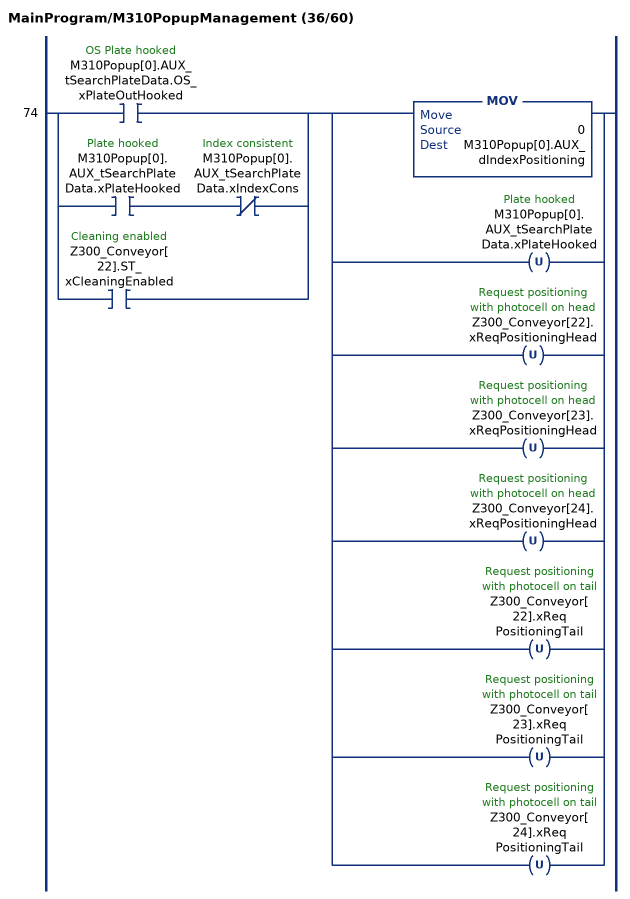
   74: [XIC(M310Popup[0].AUX_tSearchPlateData.OS_xPlateOutHooked) ,XIC(M310Popup[0].AUX_tSearchPlateData.xPlateHooked) XIO(M310Popup[0].AUX_tSearchPlateData.xIndexCons) ,XIC(Z300_Conveyor[22].ST_xCleaningEnabled) ][MOV(0,M310Popup[0].AUX_dIndexPositioning) ,OTU(M310Popup[0].AUX_tSearchPlateData.xPlateHooked) ,OTU(Z300_Conveyor[22].xReqPositioningHead) ,OTU(Z300_Conveyor[23].xReqPositioningHead) ,OTU(Z300_Conveyor[24].xReqPositioningHead) ,OTU(Z300_Conveyor[22].xReqPositioningTail) ,OTU(Z300_Conveyor[23].xReqPositioningTail) ,OTU(Z300_Conveyor[24].xReqPositioningTail) ];
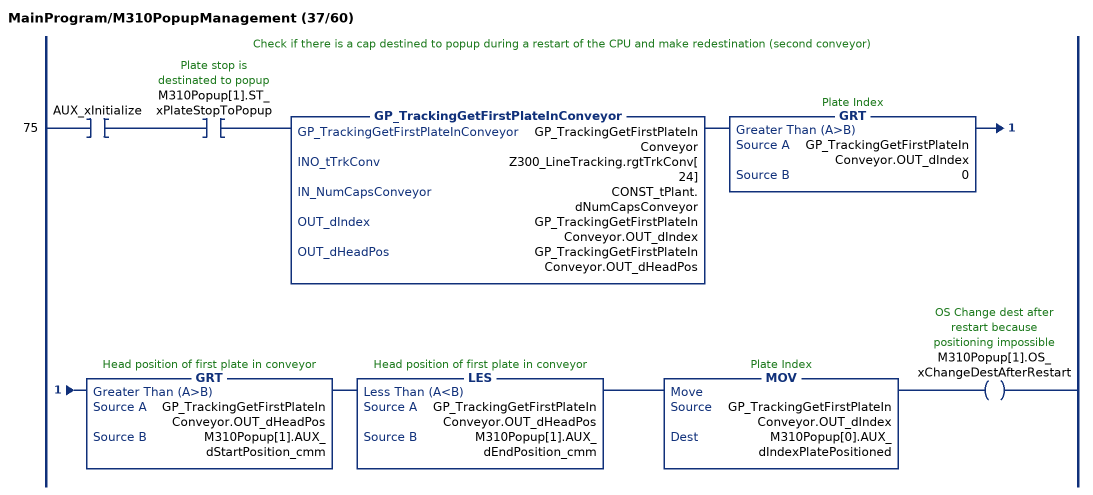
   // Check if there is a cap destined to popup during a restart of the CPU and make redestination (second conveyor)
   75: XIC(AUX_xInitialize)XIC(M310Popup[1].ST_xPlateStopToPopup)GP_TrackingGetFirstPlateInConveyor(GP_TrackingGetFirstPlateInConveyor,Z300_LineTracking.rgtTrkConv[24],CONST_tPlant.dNumCapsConveyor,GP_TrackingGetFirstPlateInConveyor.OUT_dIndex,GP_TrackingGetFirstPlateInConveyor.OUT_dHeadPos)GRT(GP_TrackingGetFirstPlateInConveyor.OUT_dIndex,0)GRT(GP_TrackingGetFirstPlateInConveyor.OUT_dHeadPos,M310Popup[1].AUX_dStartPosition_cmm)LES(GP_TrackingGetFirstPlateInConveyor.OUT_dHeadPos,M310Popup[1].AUX_dEndPosition_cmm)MOV(GP_TrackingGetFirstPlateInConveyor.OUT_dIndex,M310Popup[0].AUX_dIndexPlatePositioned)OTE(M310Popup[1].OS_xChangeDestAfterRestart);
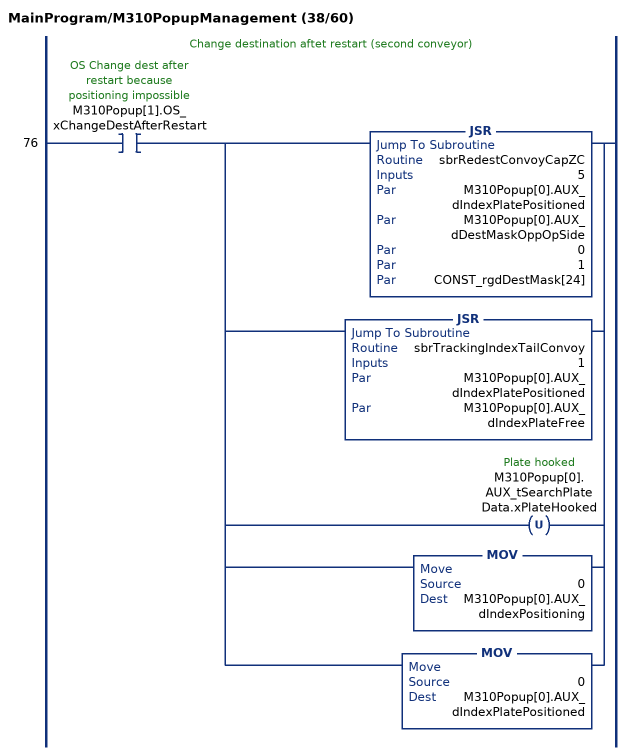
   // Change destination aftet restart (second conveyor)
   76: XIC(M310Popup[1].OS_xChangeDestAfterRestart)[JSR(sbrRedestConvoyCapZC,5,M310Popup[0].AUX_dIndexPlatePositioned,M310Popup[0].AUX_dDestMaskOppOpSide,0,1,CONST_rgdDestMask[24]) ,JSR(sbrTrackingIndexTailConvoy,1,M310Popup[0].AUX_dIndexPlatePositioned,M310Popup[0].AUX_dIndexPlateFree) ,OTU(M310Popup[0].AUX_tSearchPlateData.xPlateHooked) ,MOV(0,M310Popup[0].AUX_dIndexPositioning) ,MOV(0,M310Popup[0].AUX_dIndexPlatePositioned) ];
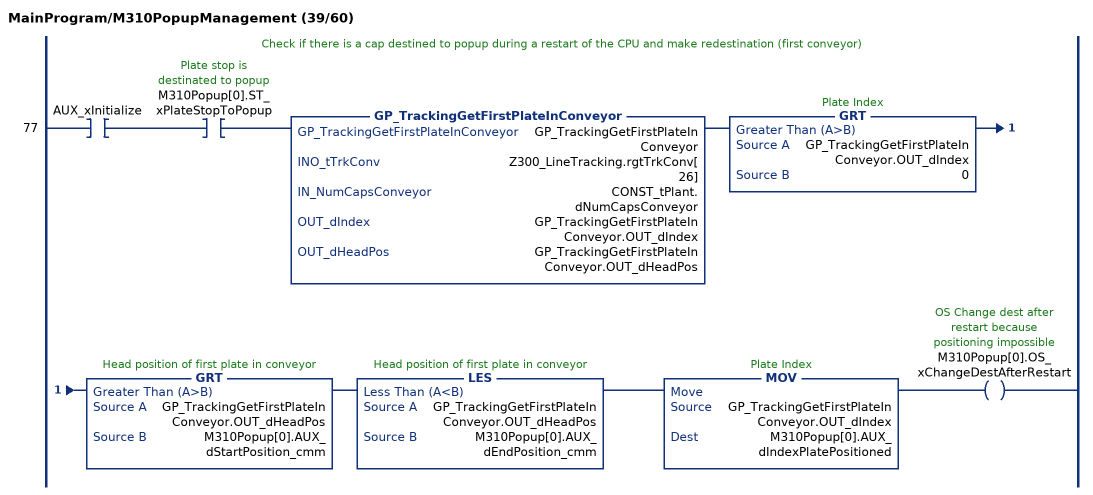
   // Check if there is a cap destined to popup during a restart of the CPU and make redestination (first conveyor)
   77: XIC(AUX_xInitialize)XIC(M310Popup[0].ST_xPlateStopToPopup)GP_TrackingGetFirstPlateInConveyor(GP_TrackingGetFirstPlateInConveyor,Z300_LineTracking.rgtTrkConv[26],CONST_tPlant.dNumCapsConveyor,GP_TrackingGetFirstPlateInConveyor.OUT_dIndex,GP_TrackingGetFirstPlateInConveyor.OUT_dHeadPos)GRT(GP_TrackingGetFirstPlateInConveyor.OUT_dIndex,0)GRT(GP_TrackingGetFirstPlateInConveyor.OUT_dHeadPos,M310Popup[0].AUX_dStartPosition_cmm)LES(GP_TrackingGetFirstPlateInConveyor.OUT_dHeadPos,M310Popup[0].AUX_dEndPosition_cmm)MOV(GP_TrackingGetFirstPlateInConveyor.OUT_dIndex,M310Popup[0].AUX_dIndexPlatePositioned)OTE(M310Popup[0].OS_xChangeDestAfterRestart);
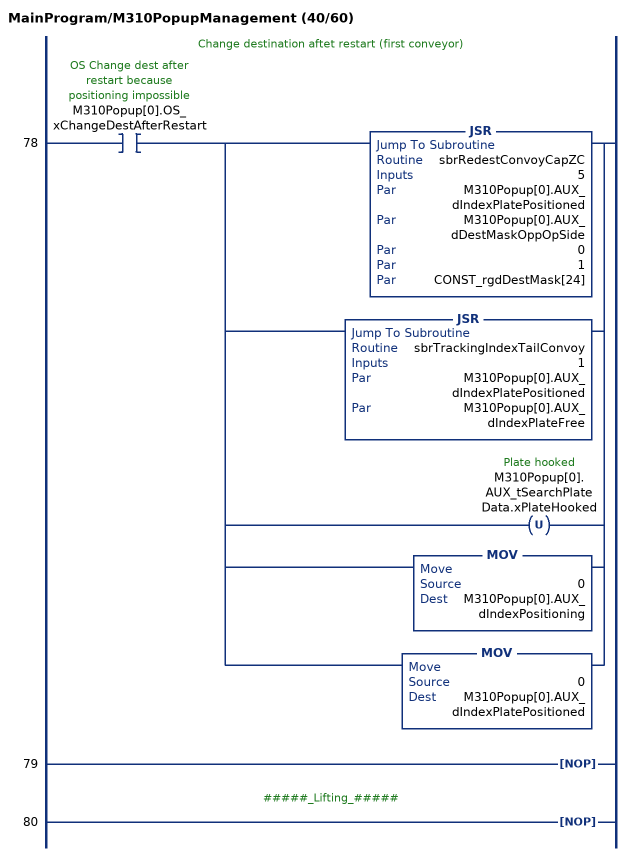
   // Change destination aftet restart (first conveyor)
   78: XIC(M310Popup[0].OS_xChangeDestAfterRestart)[JSR(sbrRedestConvoyCapZC,5,M310Popup[0].AUX_dIndexPlatePositioned,M310Popup[0].AUX_dDestMaskOppOpSide,0,1,CONST_rgdDestMask[24]) ,JSR(sbrTrackingIndexTailConvoy,1,M310Popup[0].AUX_dIndexPlatePositioned,M310Popup[0].AUX_dIndexPlateFree) ,OTU(M310Popup[0].AUX_tSearchPlateData.xPlateHooked) ,MOV(0,M310Popup[0].AUX_dIndexPositioning) ,MOV(0,M310Popup[0].AUX_dIndexPlatePositioned) ];
   79: NOP();
   // #####_Lifting_#####
   80: NOP();
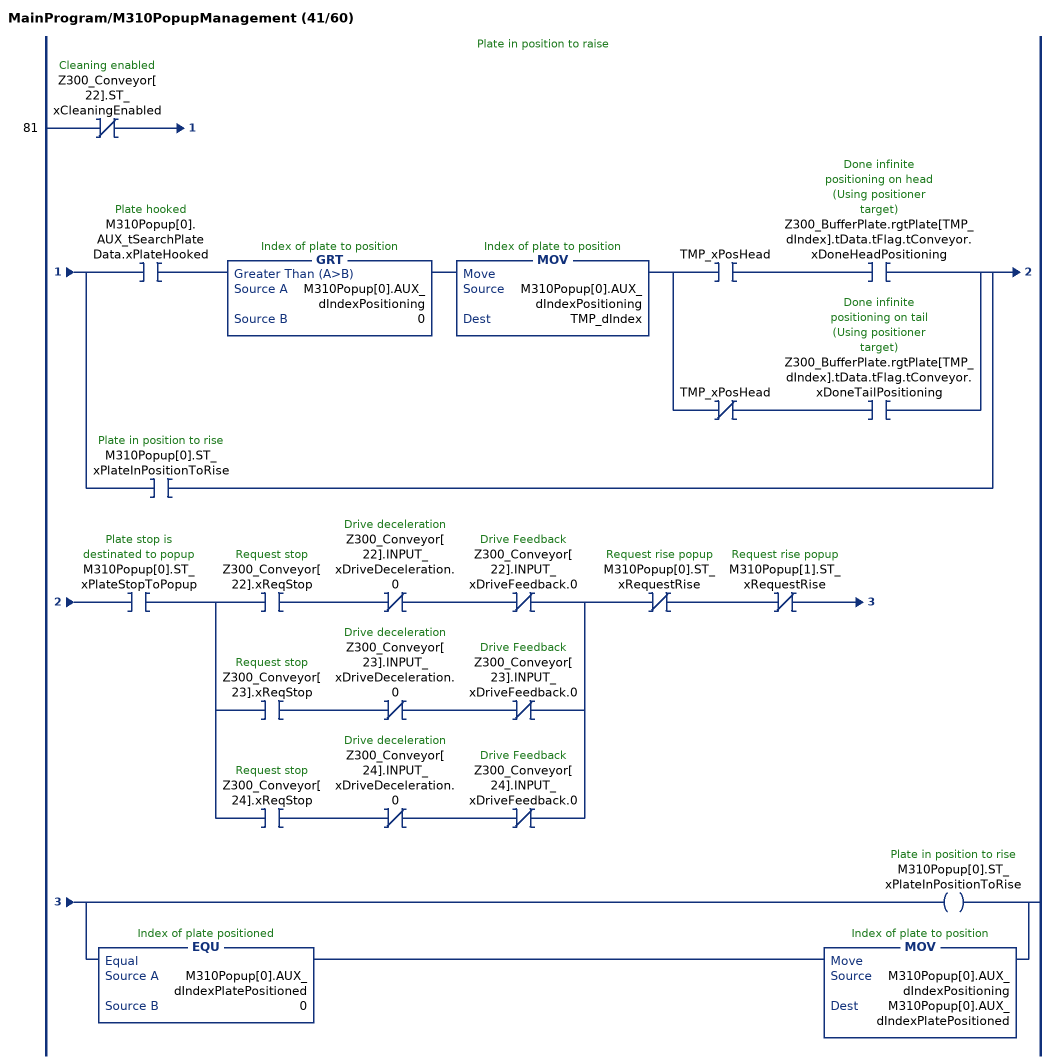
   // Plate in position to raise
   81: XIO(Z300_Conveyor[22].ST_xCleaningEnabled)[XIC(M310Popup[0].AUX_tSearchPlateData.xPlateHooked) GRT(M310Popup[0].AUX_dIndexPositioning,0) MOV(M310Popup[0].AUX_dIndexPositioning,TMP_dIndex) [XIC(TMP_xPosHead) XIC(Z300_BufferPlate.rgtPlate[TMP_dIndex].tData.tFlag.tConveyor.xDoneHeadPositioning) ,XIO(TMP_xPosHead) XIC(Z300_BufferPlate.rgtPlate[TMP_dIndex].tData.tFlag.tConveyor.xDoneTailPositioning) ] ,XIC(M310Popup[0].ST_xPlateInPositionToRise) ]XIC(M310Popup[0].ST_xPlateStopToPopup)[XIC(Z300_Conveyor[22].xReqStop) XIO(Z300_Conveyor[22].INPUT_xDriveDeceleration.0) XIO(Z300_Conveyor[22].INPUT_xDriveFeedback.0) ,XIC(Z300_Conveyor[23].xReqStop) XIO(Z300_Conveyor[23].INPUT_xDriveDeceleration.0) XIO(Z300_Conveyor[23].INPUT_xDriveFeedback.0) ,XIC(Z300_Conveyor[24].xReqStop) XIO(Z300_Conveyor[24].INPUT_xDriveDeceleration.0) XIO(Z300_Conveyor[24].INPUT_xDriveFeedback.0) ]XIO(M310Popup[0].ST_xRequestRise)XIO(M310Popup[1].ST_xRequestRise)[OTE(M310Popup[0].ST_xPlateInPositionToRise) ,EQU(M310Popup[0].AUX_dIndexPlatePositioned,0) MOV(M310Popup[0].AUX_dIndexPositioning,M310Popup[0].AUX_dIndexPlatePositioned) ];
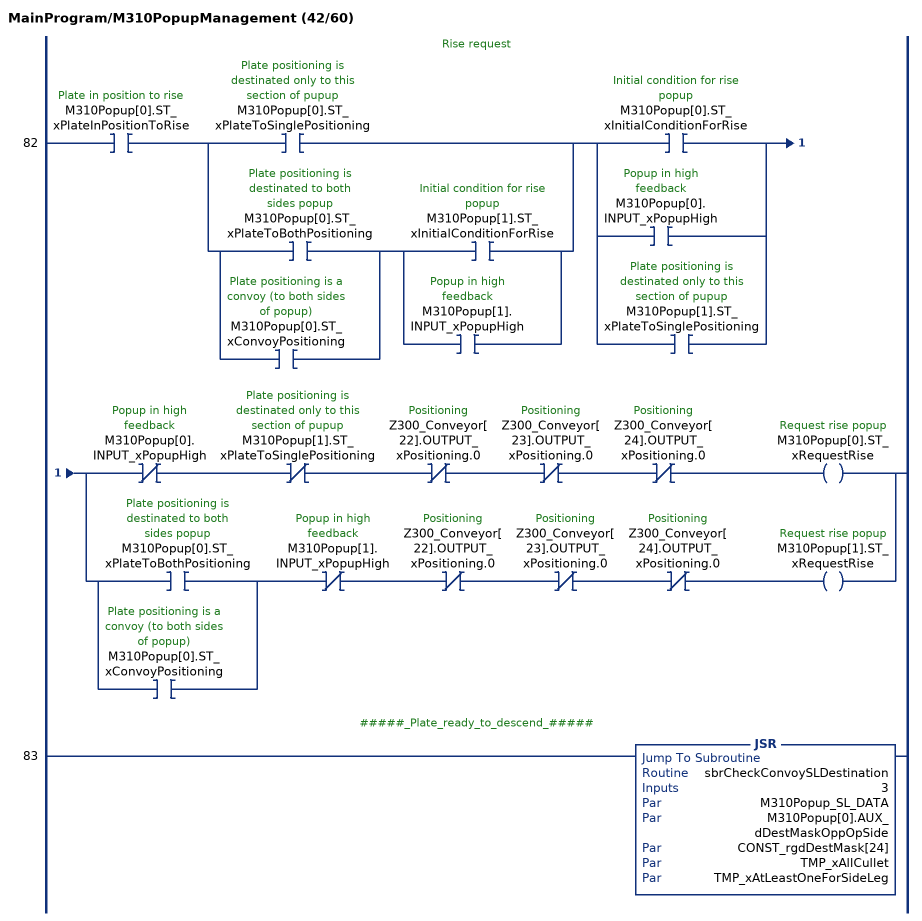
   // Rise request
   82: XIC(M310Popup[0].ST_xPlateInPositionToRise)[XIC(M310Popup[0].ST_xPlateToSinglePositioning) ,[XIC(M310Popup[0].ST_xPlateToBothPositioning) ,XIC(M310Popup[0].ST_xConvoyPositioning) ] [XIC(M310Popup[1].ST_xInitialConditionForRise) ,XIC(M310Popup[1].INPUT_xPopupHigh) ] ][XIC(M310Popup[0].ST_xInitialConditionForRise) ,XIC(M310Popup[0].INPUT_xPopupHigh) ,XIC(M310Popup[1].ST_xPlateToSinglePositioning) ][XIO(M310Popup[0].INPUT_xPopupHigh) XIO(M310Popup[1].ST_xPlateToSinglePositioning) XIO(Z300_Conveyor[22].OUTPUT_xPositioning.0) XIO(Z300_Conveyor[23].OUTPUT_xPositioning.0) XIO(Z300_Conveyor[24].OUTPUT_xPositioning.0) OTE(M310Popup[0].ST_xRequestRise) ,[XIC(M310Popup[0].ST_xPlateToBothPositioning) ,XIC(M310Popup[0].ST_xConvoyPositioning) ] XIO(M310Popup[1].INPUT_xPopupHigh) XIO(Z300_Conveyor[22].OUTPUT_xPositioning.0) XIO(Z300_Conveyor[23].OUTPUT_xPositioning.0) XIO(Z300_Conveyor[24].OUTPUT_xPositioning.0) OTE(M310Popup[1].ST_xRequestRise) ];
   // #####_Plate_ready_to_descend_#####
   83: JSR(sbrCheckConvoySLDestination,3,M310Popup_SL_DATA,M310Popup[0].AUX_dDestMaskOppOpSide,CONST_rgdDestMask[24],TMP_xAllCullet,TMP_xAtLeastOneForSideLeg);
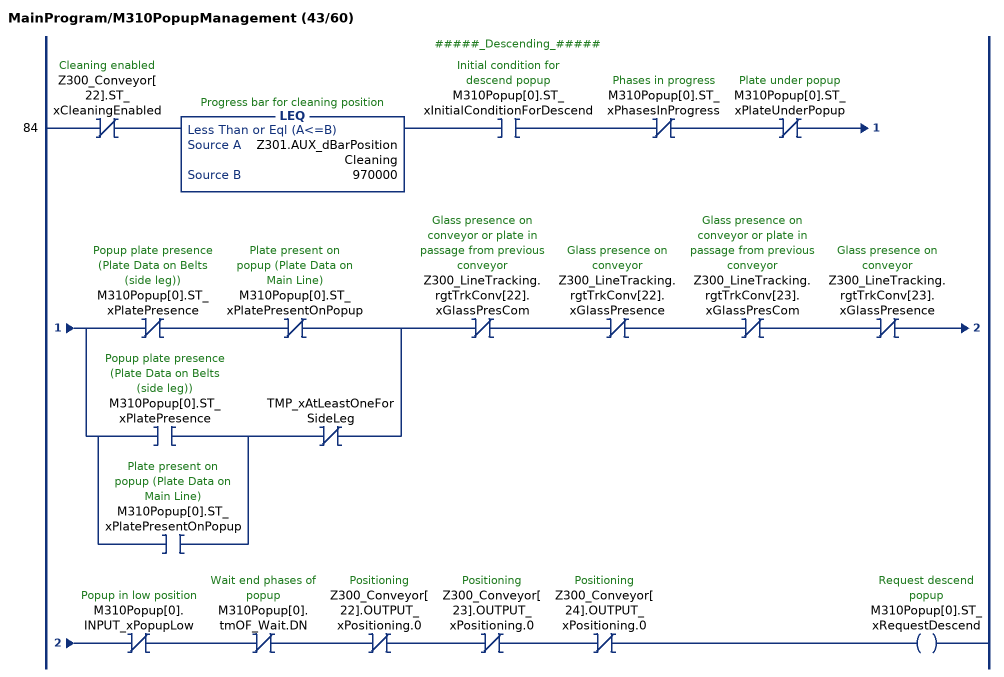
   // #####_Descending_#####
   84: XIO(Z300_Conveyor[22].ST_xCleaningEnabled)LEQ(Z301.AUX_dBarPositionCleaning,970000)XIC(M310Popup[0].ST_xInitialConditionForDescend)XIO(M310Popup[0].ST_xPhasesInProgress)XIO(M310Popup[0].ST_xPlateUnderPopup)[XIO(M310Popup[0].ST_xPlatePresence) XIO(M310Popup[0].ST_xPlatePresentOnPopup) ,[XIC(M310Popup[0].ST_xPlatePresence) ,XIC(M310Popup[0].ST_xPlatePresentOnPopup) ] XIO(TMP_xAtLeastOneForSideLeg) ]XIO(Z300_LineTracking.rgtTrkConv[22].xGlassPresCom)XIO(Z300_LineTracking.rgtTrkConv[22].xGlassPresence)XIO(Z300_LineTracking.rgtTrkConv[23].xGlassPresCom)XIO(Z300_LineTracking.rgtTrkConv[23].xGlassPresence)XIO(M310Popup[0].INPUT_xPopupLow)XIO(M310Popup[0].tmOF_Wait.DN)XIO(Z300_Conveyor[22].OUTPUT_xPositioning.0)XIO(Z300_Conveyor[23].OUTPUT_xPositioning.0)XIO(Z300_Conveyor[24].OUTPUT_xPositioning.0)OTE(M310Popup[0].ST_xRequestDescend);
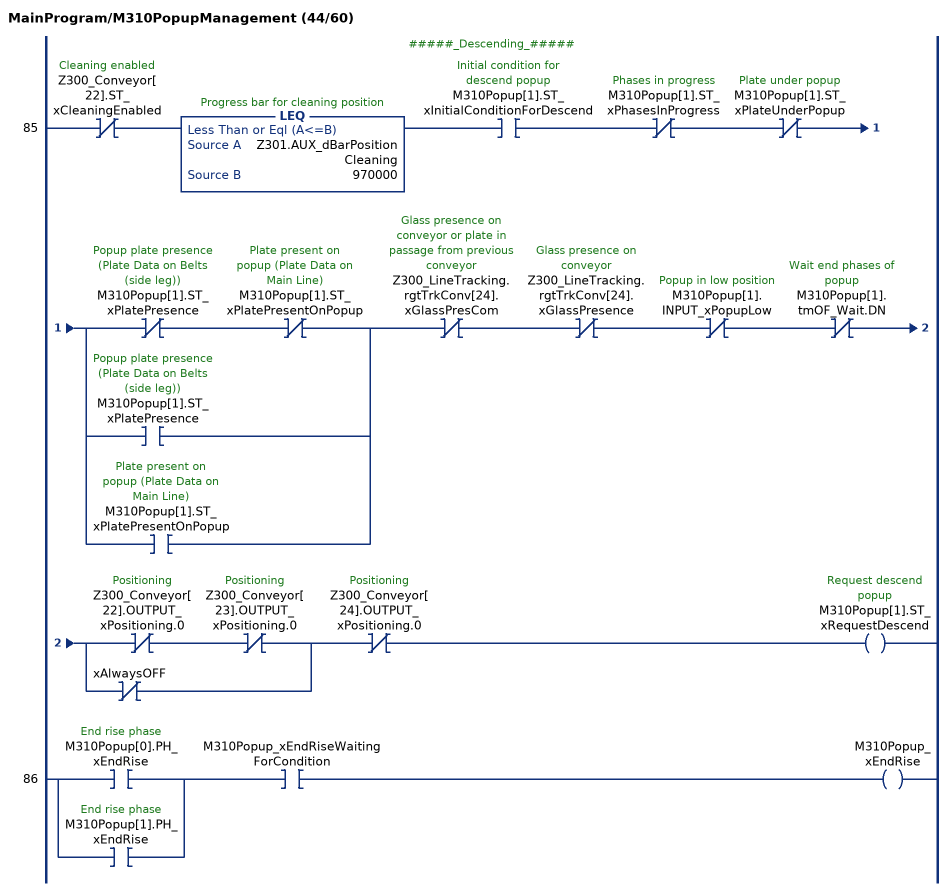
   // #####_Descending_#####
   85: XIO(Z300_Conveyor[22].ST_xCleaningEnabled)LEQ(Z301.AUX_dBarPositionCleaning,970000)XIC(M310Popup[1].ST_xInitialConditionForDescend)XIO(M310Popup[1].ST_xPhasesInProgress)XIO(M310Popup[1].ST_xPlateUnderPopup)[XIO(M310Popup[1].ST_xPlatePresence) XIO(M310Popup[1].ST_xPlatePresentOnPopup) ,[XIC(M310Popup[1].ST_xPlatePresence) ,XIC(M310Popup[1].ST_xPlatePresentOnPopup) ] ]XIO(Z300_LineTracking.rgtTrkConv[24].xGlassPresCom)XIO(Z300_LineTracking.rgtTrkConv[24].xGlassPresence)XIO(M310Popup[1].INPUT_xPopupLow)XIO(M310Popup[1].tmOF_Wait.DN)[XIO(Z300_Conveyor[22].OUTPUT_xPositioning.0) XIO(Z300_Conveyor[23].OUTPUT_xPositioning.0) ,XIO(xAlwaysOFF) ]XIO(Z300_Conveyor[24].OUTPUT_xPositioning.0)OTE(M310Popup[1].ST_xRequestDescend);
   86: [XIC(M310Popup[0].PH_xEndRise) ,XIC(M310Popup[1].PH_xEndRise) ]XIC(M310Popup_xEndRiseWaitingForCondition)OTE(M310Popup_xEndRise);
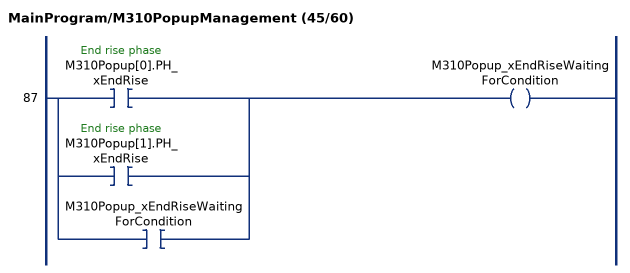
   87: [XIC(M310Popup[0].PH_xEndRise) ,XIC(M310Popup[1].PH_xEndRise) ,XIC(M310Popup_xEndRiseWaitingForCondition) ]OTE(M310Popup_xEndRiseWaitingForCondition);
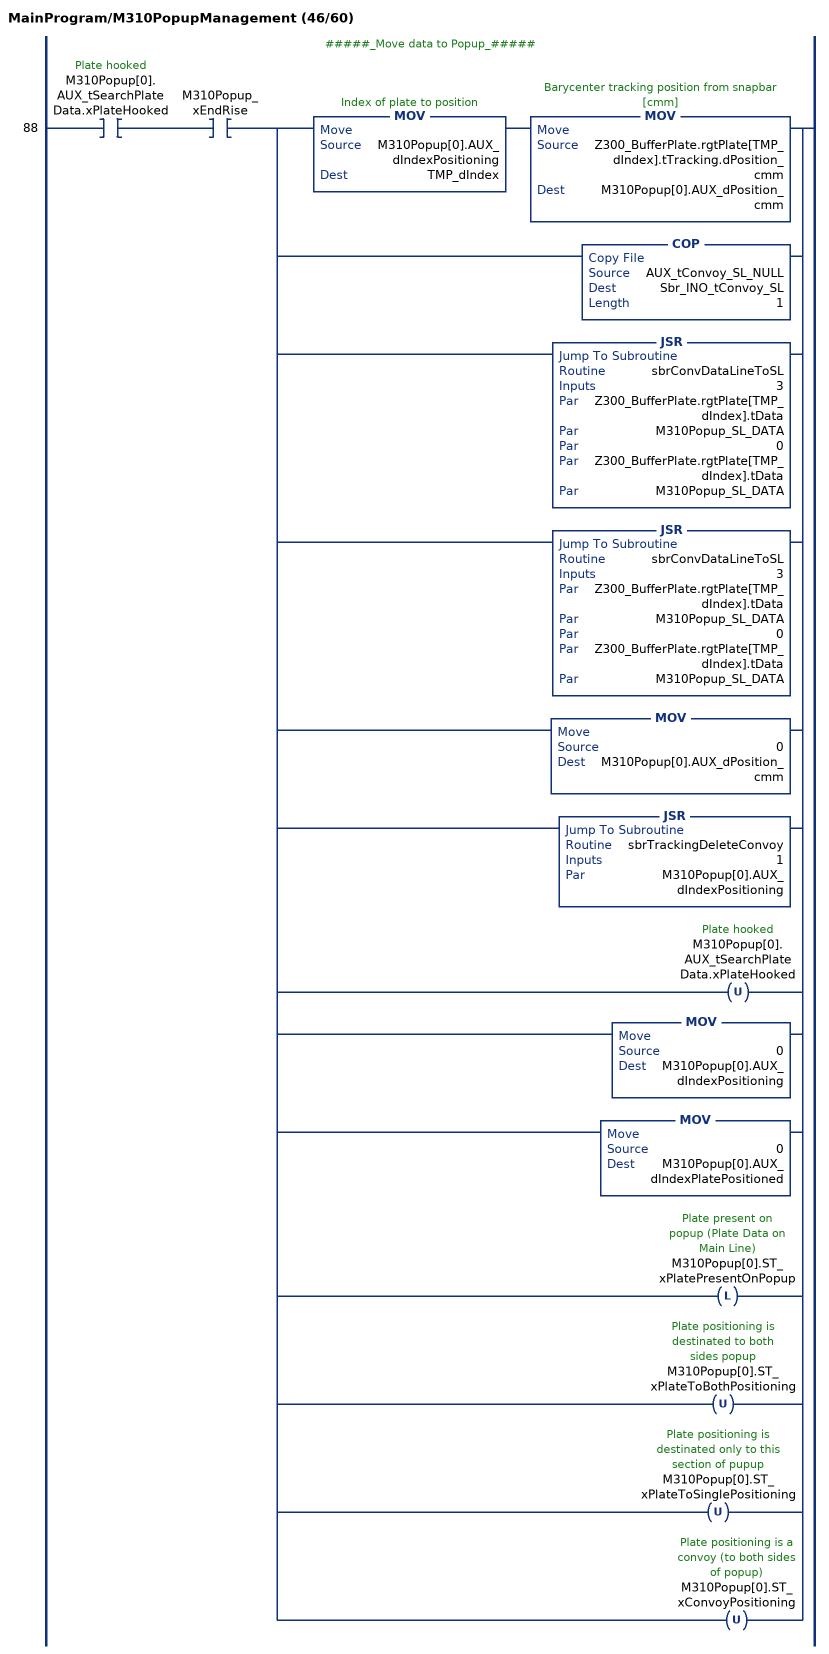
   // #####_Move data to Popup_#####
   88: XIC(M310Popup[0].AUX_tSearchPlateData.xPlateHooked)XIC(M310Popup_xEndRise)[MOV(M310Popup[0].AUX_dIndexPositioning,TMP_dIndex) MOV(Z300_BufferPlate.rgtPlate[TMP_dIndex].tTracking.dPosition_cmm,M310Popup[0].AUX_dPosition_cmm) ,COP(AUX_tConvoy_SL_NULL,Sbr_INO_tConvoy_SL,1) ,JSR(sbrConvDataLineToSL,3,Z300_BufferPlate.rgtPlate[TMP_dIndex].tData,M310Popup_SL_DATA,0,Z300_BufferPlate.rgtPlate[TMP_dIndex].tData,M310Popup_SL_DATA) ,JSR(sbrConvDataLineToSL,3,Z300_BufferPlate.rgtPlate[TMP_dIndex].tData,M310Popup_SL_DATA,0,Z300_BufferPlate.rgtPlate[TMP_dIndex].tData,M310Popup_SL_DATA) ,MOV(0,M310Popup[0].AUX_dPosition_cmm) ,JSR(sbrTrackingDeleteConvoy,1,M310Popup[0].AUX_dIndexPositioning) ,OTU(M310Popup[0].AUX_tSearchPlateData.xPlateHooked) ,MOV(0,M310Popup[0].AUX_dIndexPositioning) ,MOV(0,M310Popup[0].AUX_dIndexPlatePositioned) ,OTL(M310Popup[0].ST_xPlatePresentOnPopup) ,OTU(M310Popup[0].ST_xPlateToBothPositioning) ,OTU(M310Popup[0].ST_xPlateToSinglePositioning) ,OTU(M310Popup[0].ST_xConvoyPositioning) ];
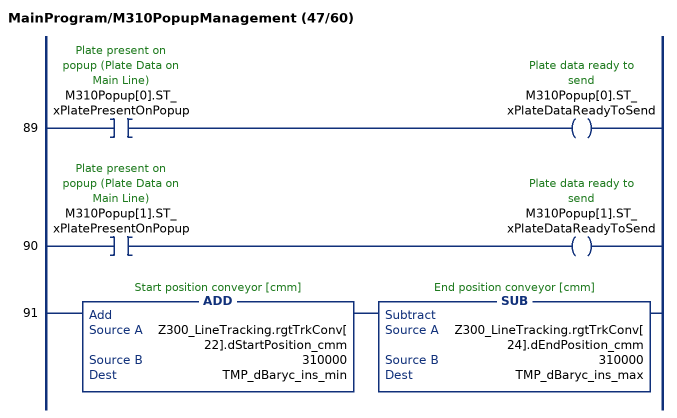
   89: XIC(M310Popup[0].ST_xPlatePresentOnPopup)OTE(M310Popup[0].ST_xPlateDataReadyToSend);
   90: XIC(M310Popup[1].ST_xPlatePresentOnPopup)OTE(M310Popup[1].ST_xPlateDataReadyToSend);
   91: ADD(Z300_LineTracking.rgtTrkConv[22].dStartPosition_cmm,310000,TMP_dBaryc_ins_min)SUB(Z300_LineTracking.rgtTrkConv[24].dEndPosition_cmm,310000,TMP_dBaryc_ins_max);
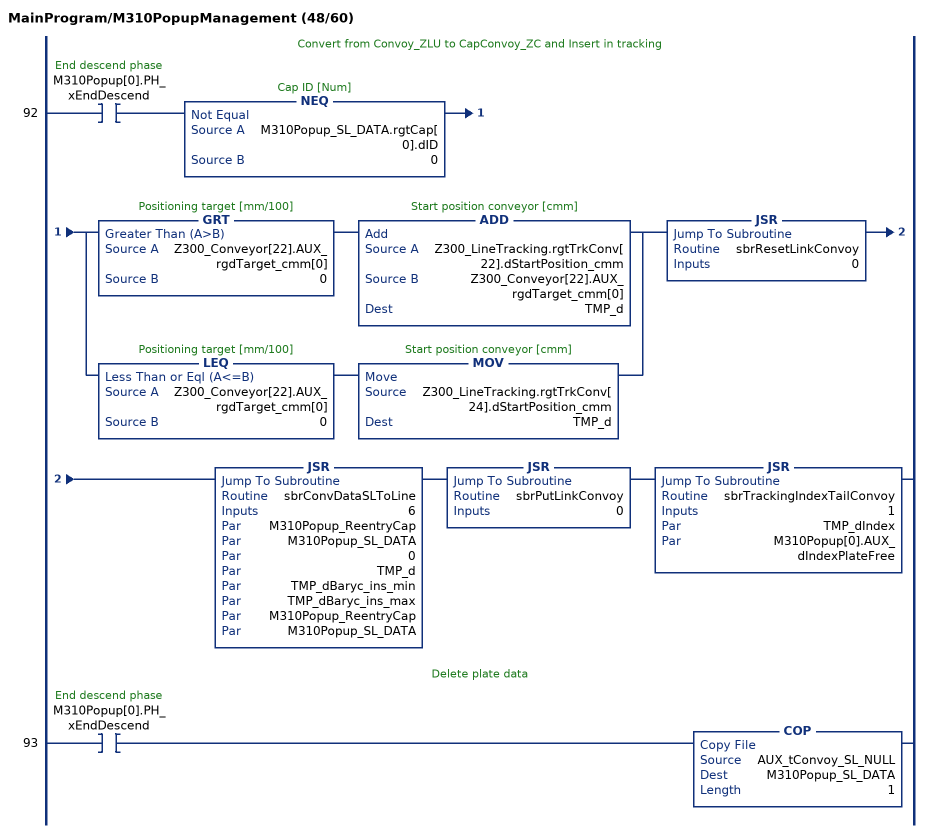
   // Convert from Convoy_ZLU to CapConvoy_ZC and Insert in tracking
   92: XIC(M310Popup[0].PH_xEndDescend)NEQ(M310Popup_SL_DATA.rgtCap[0].dID,0)[GRT(Z300_Conveyor[22].AUX_rgdTarget_cmm[0],0) ADD(Z300_LineTracking.rgtTrkConv[22].dStartPosition_cmm,Z300_Conveyor[22].AUX_rgdTarget_cmm[0],TMP_d) ,LEQ(Z300_Conveyor[22].AUX_rgdTarget_cmm[0],0) MOV(Z300_LineTracking.rgtTrkConv[24].dStartPosition_cmm,TMP_d) ]JSR(sbrResetLinkConvoy,0)JSR(sbrConvDataSLToLine,6,M310Popup_ReentryCap,M310Popup_SL_DATA,0,TMP_d,TMP_dBaryc_ins_min,TMP_dBaryc_ins_max,M310Popup_ReentryCap,M310Popup_SL_DATA)JSR(sbrPutLinkConvoy,0)JSR(sbrTrackingIndexTailConvoy,1,TMP_dIndex,M310Popup[0].AUX_dIndexPlateFree);
   // Delete plate data
   93: XIC(M310Popup[0].PH_xEndDescend)COP(AUX_tConvoy_SL_NULL,M310Popup_SL_DATA,1);
